(* Logix 5000 project; controller PLC_MCC1300_75F1 vendor 1 type 14 code 166 rev 32.11; software revision 32.04; part 62 of 83 *)
(* tags used below, declared in another part *)
   CONST_rgdDestMask : DINT[32];   // Destination Mask
   CONST_tPlant : UDT_PLANT_CONSTANTS;
   GP_TrackingSearchPlate : GP_TrackingSearchPlate;
   GP_TrackingValidateIndex : GP_TrackingValidateIndex;
   M315_M1_DR_R1 : AXIS_CIP_DRIVE;
   M315_xReqStopPrevConvForPos : BOOL;
   M315Popup : MAC_Popup_ZC[2];
   M315Popup_HMR : MAC_Popup_ZC_HMR[2];
   M315Popup_HMW : MAC_Popup_ZC_HMW[2];
   M315Popup_PlateFreeTimeout : TIMER;
   M315Popup_xDrivePosEnable : BOOL;
   TMP_d : DINT;
   TMP_dDiffPhotocellStartConv0 : DINT;
   TMP_dEndSearch0 : DINT;
   TMP_dEndSearch1 : DINT;
   TMP_dFixedSideOffsetBoth : DINT;
   TMP_dFixedSideOffsetConvoy : DINT;
   TMP_dFixedSideOffsetDW : DINT;
   TMP_dFixedSideOffsetUP : DINT;
   TMP_dHalfConveyorLength : DINT;
   TMP_dHalfPlateLength : DINT;
   TMP_dIndex : DINT;
   TMP_dStartSearch0 : DINT;
   TMP_dStartSearch1 : DINT;
   TMP_xALLForSideLeg : BOOL;
   TMP_xAllLiteToCullet : BOOL;
   TMP_xAtLeastOneForSideLeg : BOOL;
   TMP_xAtLeastOneToCullet : BOOL;
   TMP_xPosHead : BOOL;
   xAlwaysOFF : BOOL;
   xAlwaysON : BOOL;
   xDebugOFF : BOOL;
   Z300_BufferPlate : UDT_LINE_BUFFER_PLATE;
   Z300_Conveyor : UDT_StandConv[29];
   Z300_Conveyor_IN_MOTION : MAC_Conveyor_ZC_IN_MOTION[29];
   Z300_Conveyor_OUT_MOTION : MAC_Conveyor_ZC_OUT_MOTION[29];
   Z300_LineTracking : UDT_LINE_TRACKING;
   Z301 : MAC_Zone_ML;
(* MainProgram, continued *)

ROUTINE M315Popup1_Logic   (* ladder *)
   // #####_CONSTANTS_#####
   0: NOP();
   1: XIC(xAlwaysON)OTE(M315Popup[1].ST_xTunnelType);
   2: DIV(Z300_LineTracking.rgtTrkConv[28].dLengthConveyor,2,TMP_dHalfConveyorLength);
   3: MOV(Z300_LineTracking.rgtTrkConv[28].dStartPosition_cmm,M315Popup[1].AUX_dStartPosition_cmm)MOV(Z300_LineTracking.rgtTrkConv[28].dEndPosition_cmm,M315Popup[1].AUX_dEndPosition_cmm)MOV(1500,M315Popup[1].AUX_dReactionTime_ms)MOV(200000,M315Popup[1].AUX_dWindowSearch_cmm)MOV(Z300_Conveyor[28].AUX_rgdCurrentSpeed_mm_min[0],M315Popup[1].AUX_dSpeedConveyor_mm_min);
   // #####_MATCH_#####
   4: NOP();
   5: XIC(Z301.ST_xEnableControlError)OTE(M315Popup[1].ST_xEnableControlError);
   // #####_ALARMS_#####
   6: NOP();
   7: JSR(M315Popup1_Faults,0);
   // #####_HMI_LOGICS_#####
   8: NOP();
   9: XIC(xAlwaysON)OTE(M315Popup[1].ST_xExternalConditionToRise);
   10: XIC(xAlwaysON)OTE(M315Popup[1].ST_xExternalConditionToDescend);
   // #####_STATUSES_#####
   11: NOP();
   12: [XIC(M315Popup[1].ST_xStopMachineFault) ,XIC(M315Popup[1].ST_xStopNextCycleFault) ]OTE(M315Popup[1].ST_xMachineAlarm);
   13: [XIO(M315Popup[1].ST_xPhasesInProgress) ,XIO(M315Popup[1].ST_xOutputEnable) ]OTE(M315Popup[1].ST_xConditionOKForStopCycle);
   14: XIC(Z301.ST_xCycleON)XIO(M315Popup[1].ST_xManualMode)XIO(M315Popup[1].ST_xMachineAlarm)OTE(M315Popup[1].ST_xOutputEnable);
   15: XIC(Z301.ST_xCycleON)XIC(M315Popup[1].ST_xOutputEnable)XIO(M315Popup[1].ST_xPhasesInProgress)XIO(M315Popup[1].INPUT_xPopupHigh)XIC(M315Popup[1].INPUT_xPopupLow)XIO(M315Popup[1].ST_xCleaningAccepted)OTE(M315Popup[1].ST_xInitialConditionForRise);
   16: XIC(Z301.ST_xCycleON)XIC(M315Popup[1].ST_xOutputEnable)XIO(M315Popup[1].ST_xPhasesInProgress)XIO(M315Popup[1].INPUT_xPopupLow)XIC(M315Popup[1].INPUT_xPopupHigh)XIO(M315Popup[1].ST_xCleaningAccepted)OTE(M315Popup[1].ST_xInitialConditionForDescend);
   17: [XIC(M315Popup_HMW[1].xEnableDisableManualCommand) XIC(xAlwaysOFF) ,XIC(Z300_Conveyor[23].ST_xManualCmdEnabled) ]XIC(M315Popup[1].ST_xConditionOKForStopCycle)XIC(M315Popup[1].ST_xConditionOKForStopCycle)OTE(M315Popup[1].ST_xManualMode);
   18: XIO(M315Popup[1].ST_xManualMode)MOV(0,M315Popup_HMW[1].rgxMan);
   // #####_PHASES_&_LOGICS_#####
   19: NOP();
   20: XIC(xAlwaysON)OTE(M315Popup[1].ST_xCleaningConditionOK);
   21: [XIC(M315Popup_HMW[1].xLocalCleaningRequest) XIC(xAlwaysOFF) ,XIC(Z300_Conveyor[28].ST_xCleaningEnabled) XIC(M315Popup[1].INPUT_xPopupLow) ][XIC(M315Popup[1].ST_xCleaningConditionOK) ,XIC(M315Popup[1].ST_xCleaningAccepted) ]OTE(M315Popup[1].ST_xCleaningAccepted);
   22: XIC(M315Popup[1].ST_xInitialConditionForRise)XIC(M315Popup[1].ST_xExternalConditionToRise)XIC(M315Popup[1].ST_xRequestRise)XIO(M315Popup[1].PH_xRise)OTL(M315Popup[1].PH_xRise);
   23: XIC(M315Popup[1].PH_xRise)XIC(M315Popup[1].INPUT_xPopupHigh)XIO(M315Popup[1].INPUT_xPopupLow)[OTU(M315Popup[1].PH_xRise) ,OTE(M315Popup[1].PH_xEndRise) ];
   24: XIC(M315Popup[1].ST_xInitialConditionForDescend)XIC(M315Popup[1].ST_xExternalConditionToDescend)XIC(M315Popup[1].ST_xRequestDescend)[XIC(M315Popup[0].ST_xRequestDescend) ,XIC(M315Popup[0].INPUT_xPopupLow) ]XIO(M315Popup[1].PH_xDescend)OTL(M315Popup[1].PH_xDescend);
   25: XIC(M315Popup[1].PH_xDescend)XIC(M315Popup[1].INPUT_xPopupLow)XIO(M315Popup[1].INPUT_xPopupHigh)[OTU(M315Popup[1].PH_xDescend) ,OTE(M315Popup[1].PH_xEndDescend) ];
   26: [XIC(M315Popup[1].PH_xRise) ,XIC(M315Popup[1].PH_xEndRise) ,XIC(M315Popup[1].PH_xDescend) ,XIC(M315Popup[1].PH_xEndDescend) ]OTE(M315Popup[1].ST_xPhasesInProgress);
   27: [XIC(M315Popup[1].PH_xEndDescend) ,XIO(xAlwaysOFF) XIC(M315Popup[0].INPUT_xPopupLow) XIC(M315Popup[1].INPUT_xPopupLow) ]OTU(M315Popup[1].ST_xPlatePresence);
   28: XIO(M315Popup[1].ST_xPhasesInProgress)[XIC(M315Popup[1].INPUT_xPopupLow) XIO(M315Popup[1].INPUT_xPopupHigh) ,XIC(M315Popup[1].ST_xTunnelType) XIC(M315Popup[1].INPUT_xPopupHigh) XIO(M315Popup[1].INPUT_xPopupLow) ]OTE(M315Popup[1].ST_xOutOfEncumbrance);
   29: XIO(M315Popup[1].ST_xPhasesInProgress)XIO(M315Popup[1].ST_xPlatePresence)XIO(M315Popup[1].INPUT_xPopupHigh)XIC(M315Popup[1].INPUT_xPopupLow)OTE(M315Popup[1].ST_xConditionToReceiveGlass);
   30: XIO(M315Popup[1].ST_xPhasesInProgress)XIC(M315Popup[1].INPUT_xPopupHigh)XIO(M315Popup[1].INPUT_xPopupLow)OTE(M315Popup[1].ST_xConditionForUpperConveyor);
   // #####_EXTERNAL_DEVICE_#####
   31: NOP();
   // #####_HMI_STATUSES_#####
   32: NOP();
   33: XIC(M315Popup[1].INPUT_xPopupHigh)OTE(M315Popup_HMR[1].xHighPosition);
   34: XIC(M315Popup[1].INPUT_xPopupLow)OTE(M315Popup_HMR[1].xLowPosition);
   35: [MOV(1,M315Popup_HMR[1].rgdState) ,[XIC(M315Popup[1].OUTPUT_xPopupLifting) ,XIC(M315Popup[1].OUTPUT_xPopupDescent) ] MOV(3,M315Popup_HMR[1].rgdState) ,XIC(M315Popup[1].ST_xMachineWarning) MOV(5,M315Popup_HMR[1].rgdState) ,XIC(M315Popup[1].ST_xMachineAlarm) MOV(7,M315Popup_HMR[1].rgdState) ];
   36: XIC(M315Popup[1].ST_xCleaningAccepted)OTE(M315Popup_HMR[1].xPopUpCleaningEnabled);
   37: XIC(M315Popup[1].ST_xManualMode)XIC(M315Popup_HMW[1].rgxMan.0)XIC(M315Popup[1].OUTPUT_xPopupLifting)OTE(M315Popup_HMR[1].rgxMan.0);
   38: XIC(M315Popup[1].ST_xManualMode)XIC(M315Popup_HMW[1].rgxMan.1)XIC(M315Popup[1].OUTPUT_xPopupDescent)OTE(M315Popup_HMR[1].rgxMan.1);
   39: XIC(M315Popup[1].ST_xManualMode)XIC(M315Popup_HMW[1].rgxMan.8)XIC(M315Popup[1].OUTPUT_xRun)OTE(M315Popup_HMR[1].rgxMan.8);
   40: XIC(M315Popup[1].ST_xManualMode)XIC(M315Popup_HMW[1].rgxMan.9)XIC(M315Popup[1].OUTPUT_xReverse)OTE(M315Popup_HMR[1].rgxMan.9);
END_ROUTINE

ROUTINE M315PopupManagement   (* ladder *)
   // #####_CONSTANTS_#####
   0: NOP();
   1: MOV(CONST_rgdDestMask[2],M315Popup[0].AUX_dDestMaskOppOpSide)MOV(CONST_rgdDestMask[2],M315Popup[1].AUX_dDestMaskOppOpSide)MOV(20000,TMP_dFixedSideOffsetUP)MOV(-20000,TMP_dFixedSideOffsetDW)MOV(43000,TMP_dFixedSideOffsetBoth)MOV(30000,TMP_dFixedSideOffsetConvoy)MOV(380000,TMP_dHalfConveyorLength);
   // #####_MATCH_#####
   2: NOP();
   3: MOV(Z300_LineTracking.rgtTrkConv[26].dStartPosition_cmm,M315Popup[0].AUX_dStartPosition_cmm)MOV(Z300_LineTracking.rgtTrkConv[27].dEndPosition_cmm,M315Popup[0].AUX_dEndPosition_cmm)MOV(M315Popup[0].AUX_dEndPosition_cmm,M315Popup[1].AUX_dStartPosition_cmm)MOV(Z300_LineTracking.rgtTrkConv[28].dEndPosition_cmm,M315Popup[1].AUX_dEndPosition_cmm);
   4: MOV(Z300_LineTracking.rgtTrkConv[26].dStartPosition_cmm,M315Popup[0].AUX_dPosPhotocell_cmm)MOV(Z300_LineTracking.rgtTrkConv[26].dStartPosition_cmm,M315Popup[1].AUX_dPosPhotocell_cmm)SUB(Z300_LineTracking.rgtTrkConv[26].dStartPosition_cmm,M315Popup[0].AUX_dPosPhotocell_cmm,TMP_dDiffPhotocellStartConv0)MOV(50,M315Popup[0].tmOF_Wait.PRE)MOV(50,M315Popup[1].tmOF_Wait.PRE)MOV(10000,M315Popup[0].tmON_Saturation.PRE)MOV(10000,M315Popup[1].tmON_Saturation.PRE);
   5: SUB(M315Popup[0].AUX_dPosPhotocell_cmm,300000,TMP_dStartSearch0)SUB(M315Popup[0].AUX_dPosPhotocell_cmm,0,TMP_dEndSearch0)SUB(M315Popup[0].AUX_dPosPhotocell_cmm,300000,TMP_dStartSearch1)SUB(M315Popup[0].AUX_dPosPhotocell_cmm,0,TMP_dEndSearch1);
   // Set Positioning Type
   6: XIC(xAlwaysON)OTE(TMP_xPosHead);
   // ##### PREVIOUS CONVEYOR #####
   7: NOP();
   // Search plate limits
   8: MUL(M315Popup[0].AUX_dSpeedConveyor_mm_min,M315Popup[0].AUX_dReactionTime_ms,TMP_d)DIV(TMP_d,600,M315Popup[0].AUX_tSearchPlateData.dReaction_cmm);
   9: MOV(TMP_dStartSearch0,M315Popup[0].AUX_tSearchPlateData.dPositionDecision_cmm)MOV(TMP_dEndSearch0,M315Popup[0].AUX_tSearchPlateData.dPositionStopSearch_cmm)ADD(Z300_LineTracking.rgtTrkConv[28].dEndPosition_cmm,300000,M315Popup[0].AUX_tSearchPlateData.dPositionStopHooked_cmm);
   // Search plate on previous conveyor (reverse search)
   10: XIO(M315Popup[0].AUX_tSearchPlateData.xPlateHooked)GP_TrackingSearchPlate(GP_TrackingSearchPlate,M315Popup[0].AUX_tSearchPlateData.dPositionStopSearch_cmm,M315Popup[0].AUX_tSearchPlateData.dPositionDecision_cmm,0,Z300_LineTracking,M315Popup[0].AUX_tSearchPlateData.tResult,CONST_tPlant.dNumOfConveyors,CONST_tPlant.dNumCapsConveyor,Z300_BufferPlate);
   11: XIO(Z300_LineTracking.rgtTrkConv[25].xGlassPresence)XIO(Z300_LineTracking.rgtTrkConv[26].xGlassPresence)XIO(Z300_LineTracking.rgtTrkConv[27].xGlassPresence)XIO(Z300_LineTracking.rgtTrkConv[28].xGlassPresence)XIC(TMP_xPosHead)XIO(M315Popup[0].AUX_tSearchPlateData.tResult.xHeadPresence)MOV(0,M315Popup[0].AUX_tSearchPlateData.dIndex)MOV(0,M315Popup[0].AUX_dIndexHead);
   12: XIO(Z300_LineTracking.rgtTrkConv[25].xGlassPresence)XIO(Z300_LineTracking.rgtTrkConv[26].xGlassPresence)XIO(Z300_LineTracking.rgtTrkConv[27].xGlassPresence)XIO(Z300_LineTracking.rgtTrkConv[28].xGlassPresence)XIO(TMP_xPosHead)XIO(M315Popup[0].AUX_tSearchPlateData.tResult.xTailPresence)MOV(0,M315Popup[0].AUX_tSearchPlateData.dIndex)MOV(0,M315Popup[0].AUX_dIndexTail);
   13: XIC(TMP_xPosHead)XIC(M315Popup[0].AUX_tSearchPlateData.tResult.xHeadPresence)MOV(M315Popup[0].AUX_tSearchPlateData.tResult.rgdHeadPointer[0],M315Popup[0].AUX_dIndexHead);
   14: XIO(TMP_xPosHead)XIC(M315Popup[0].AUX_tSearchPlateData.tResult.xTailPresence)MOV(M315Popup[0].AUX_tSearchPlateData.tResult.rgdTailPointer[0],M315Popup[0].AUX_dIndexTail);
   15: XIO(M315Popup[0].AUX_tSearchPlateData.xPlateHooked)[XIC(TMP_xPosHead) XIC(M315Popup[0].AUX_tSearchPlateData.tResult.xHeadPresence) MOV(M315Popup[0].AUX_tSearchPlateData.tResult.rgdHeadPointer[0],M315Popup[0].AUX_tSearchPlateData.dIndex) ,XIO(TMP_xPosHead) XIC(M315Popup[0].AUX_tSearchPlateData.tResult.xTailPresence) MOV(M315Popup[0].AUX_tSearchPlateData.tResult.rgdTailPointer[0],M315Popup[0].AUX_tSearchPlateData.dIndex) ][OSR(M315Popup[0].AUX_tSearchPlateData.OSR_xPlateInWindows,M315Popup[0].AUX_tSearchPlateData.OS_xPlateInWindows) ,OSF(M315Popup[0].AUX_tSearchPlateData.OSF_xPlateInWindows,M315Popup[0].AUX_tSearchPlateData.OF_xPlateInWindows) ];
   16: GRT(M315Popup[0].AUX_tSearchPlateData.dIndex,0)[OTU(TMP_xAtLeastOneForSideLeg) ,OTL(TMP_xALLForSideLeg) ,OTL(TMP_xAllLiteToCullet) ,OTU(TMP_xAtLeastOneToCullet) ];
   // Verify destination
   17: GRT(M315Popup[0].AUX_tSearchPlateData.dIndex,0)JSR(sbrCheckConvoyZCDestination,5,M315Popup[0].AUX_tSearchPlateData.dIndex,M315Popup[0].AUX_dDestMaskOppOpSide,CONST_rgdDestMask[24],TMP_xAtLeastOneForSideLeg,TMP_xAllLiteToCullet,TMP_xAtLeastOneForSideLeg,TMP_xAllLiteToCullet)JSR(sbrCheckConvoyZCDestinationFull,5,M315Popup[0].AUX_tSearchPlateData.dIndex,M315Popup[0].AUX_dDestMaskOppOpSide,CONST_rgdDestMask[24],TMP_xALLForSideLeg,TMP_xAtLeastOneToCullet,TMP_xALLForSideLeg,TMP_xAtLeastOneToCullet)[XIC(TMP_xAtLeastOneForSideLeg) XIC(TMP_xALLForSideLeg) OTE(M315Popup[0].ST_xPlateComingToPopup) ,XIO(TMP_xALLForSideLeg) MOV(M315Popup[0].AUX_tSearchPlateData.dIndex,M315Popup[0].AUX_dIndexPlateFree) ];
   18: GP_TrackingValidateIndex(GP_TrackingValidateIndex,Z300_BufferPlate,M315Popup[0].AUX_tSearchPlateData.dIDMemory,M315Popup[0].AUX_tSearchPlateData.dIndex,M315Popup[0].AUX_tSearchPlateData.xIndexCons);
   // Check plate dimension
   19: XIC(M315Popup[0].ST_xPlateComingToPopup)MOV(M315Popup[0].AUX_tSearchPlateData.dIndex,TMP_dIndex)[LEQ(Z300_BufferPlate.rgtPlate[TMP_dIndex].tData.dTotalCaps,1) [GRT(Z300_BufferPlate.rgtPlate[TMP_dIndex].tData.dLength_cmm,TMP_dHalfConveyorLength) OTE(M315Popup[0].ST_xPlateToBothComing) ,XIO(M315Popup[0].ST_xPlateToBothComing) OTE(M315Popup[0].ST_xPlateToSingleComing) ] ,GRT(Z300_BufferPlate.rgtPlate[TMP_dIndex].tData.dTotalCaps,1) [LEQ(Z300_BufferPlate.rgtPlate[TMP_dIndex].tData.dLength_cmm,CONST_tPlant.rgdConvoyLimits_cmm[2]) ,XIO(xAlwaysOFF) ] OTE(M315Popup[0].ST_xConvoyComing) ];
   20: [XIC(Z300_Conveyor[25].xReqStop) ,XIO(xAlwaysOFF) ]XIC(M315Popup[0].ST_xPhasesInProgress)TOF(M315Popup[0].tmOF_Wait,?,?);
   21: [XIC(Z300_Conveyor[25].xReqStop) ,XIO(xAlwaysOFF) ]XIC(M315Popup[1].ST_xPhasesInProgress)TOF(M315Popup[1].tmOF_Wait,?,?);
   // Plate has left popup conveyors
   22: GRT(M315Popup[0].AUX_dIndexPlateFree,0)MOV(M315Popup[0].AUX_dIndexPlateFree,TMP_dIndex)GEQ(Z300_BufferPlate.rgtPlate[TMP_dIndex].tTracking.dPositionTail_cmm,Z300_LineTracking.rgtTrkConv[24].dEndPosition_cmm)MOV(0,M315Popup[0].AUX_dIndexPlateFree);
   // Stop previuos conveyor if no condition on pop-up conveyor
   23: [[XIC(M315Popup[0].ST_xPlateToSingleComing) [XIO(M315Popup[0].ST_xInitialConditionForRise) ,XIC(M315Popup[0].ST_xPlatePresentOnPopup) ,XIC(M315Popup[0].ST_xPlatePresence) ,XIC(Z300_LineTracking.rgtTrkConv[26].xGlassPresence) ,XIC(Z300_LineTracking.rgtTrkConv[27].xGlassPresence) ,EQU(M315Popup[0].AUX_dIndexPositioning,0) [XIC(M315Popup[0].ST_xPlateUnderPopup) ,XIC(M315Popup[1].ST_xPlateUnderPopup) ] ] ,XIC(M315Popup[0].ST_xPlateToSingleComing) [XIO(M315Popup[1].ST_xInitialConditionForRise) ,XIC(M315Popup[1].ST_xPlatePresentOnPopup) ,XIC(M315Popup[1].ST_xPlatePresence) ,XIC(Z300_LineTracking.rgtTrkConv[26].xGlassPresence) ,XIC(Z300_LineTracking.rgtTrkConv[27].xGlassPresence) ,XIC(Z300_LineTracking.rgtTrkConv[28].xGlassPresence) ,EQU(M315Popup[0].AUX_dIndexPositioning,0) [XIC(M315Popup[0].ST_xPlateUnderPopup) ,XIC(M315Popup[1].ST_xPlateUnderPopup) ] ] ,[XIC(M315Popup[0].ST_xPlateToBothComing) ,XIC(M315Popup[0].ST_xConvoyComing) ] [XIO(M315Popup[1].ST_xInitialConditionForRise) ,XIC(M315Popup[1].ST_xPlatePresentOnPopup) ,XIC(M315Popup[1].ST_xPlatePresence) ,XIC(Z300_LineTracking.rgtTrkConv[26].xGlassPresence) ,XIC(Z300_LineTracking.rgtTrkConv[27].xGlassPresence) ,XIC(Z300_LineTracking.rgtTrkConv[28].xGlassPresence) ,EQU(M315Popup[0].AUX_dIndexPositioning,0) XIC(M315Popup[1].ST_xPlateUnderPopup) ,XIO(M315Popup[0].ST_xInitialConditionForRise) ,XIC(M315Popup[0].ST_xPlatePresentOnPopup) ,XIC(M315Popup[0].ST_xPlatePresence) ,EQU(M315Popup[0].AUX_dIndexPositioning,0) XIC(M315Popup[0].ST_xPlateUnderPopup) ] ] ,XIO(M315Popup[0].INPUT_xPopupHigh) XIO(M315Popup[0].INPUT_xPopupLow) ,XIO(M315Popup[1].INPUT_xPopupHigh) XIO(M315Popup[1].INPUT_xPopupLow) ,XIC(M315_xReqStopPrevConvForPos) ,XIC(Z300_Conveyor[26].xReqExtStopLoadNewPlate) ,[XIC(M315Popup[0].ST_xPlateInPositionToRise) ,XIC(M315Popup[1].ST_xPlateInPositionToRise) ] ,XIC(Z300_Conveyor[26].ST_xCleaningEnabled) XIO(Z300_Conveyor[25].ST_xCleaningEnabled) ,XIC(M315Popup[0].ST_xPrevConvFreeAfterPos) ,XIC(M315Popup[1].ST_xPrevConvFreeAfterPos) ,[XIO(M315Popup[0].INPUT_xPopupHigh) ,XIO(M315Popup[1].INPUT_xPopupHigh) ] ,GRT(M315Popup[0].AUX_dIndexPositioning,0) [GRT(M315Popup[0].AUX_tSearchPlateData.dIndex,0) NEQ(M315Popup[0].AUX_tSearchPlateData.dIndex,M315Popup[0].AUX_dIndexPositioning) ,GRT(M315Popup[0].AUX_dIndexPlatePositioned,0) NEQ(M315Popup[0].AUX_dIndexPlatePositioned,M315Popup[0].AUX_dIndexPositioning) ] ,GRT(M315Popup[0].AUX_dIndexPlateFree,0) MOV(M315Popup[0].AUX_dIndexPlateFree,TMP_dIndex) [XIC(M315Popup[0].ST_xPlateToSingleComing) LES(Z300_BufferPlate.rgtPlate[TMP_dIndex].tTracking.dPositionTail_cmm,M315Popup[1].AUX_dStartPosition_cmm) ,[XIC(M315Popup[0].ST_xPlateToBothComing) ,XIC(M315Popup[0].ST_xConvoyComing) ,XIC(M315Popup[1].ST_xPlateToSingleComing) ] LES(Z300_BufferPlate.rgtPlate[TMP_dIndex].tTracking.dPositionTail_cmm,Z300_LineTracking.rgtTrkConv[24].dEndPosition_cmm) ] ]OTE(M315Popup[0].ST_xConditionToStopPrevious);
   24: XIO(xDebugOFF)GRT(M315Popup[0].AUX_dIndexPlateFree,0)XIC(Z300_Conveyor[26].ST_xRotationFeedback)MOV(10000,M315Popup_PlateFreeTimeout.PRE)[TON(M315Popup_PlateFreeTimeout,?,?) ,XIC(M315Popup_PlateFreeTimeout.DN) MOV(0,M315Popup[0].AUX_dIndexPlateFree) ];
   25: XIO(Z300_LineTracking.rgtTrkConv[26].xGlassPresence)XIO(Z300_LineTracking.rgtTrkConv[27].xGlassPresence)XIO(Z300_LineTracking.rgtTrkConv[28].xGlassPresence)XIC(Z300_Conveyor[26].ST_xRotationFeedback)XIC(Z300_Conveyor[27].ST_xRotationFeedback)XIC(Z300_Conveyor[28].ST_xRotationFeedback)[GRT(M315Popup[0].AUX_dIndexPlateFree,0) ,GRT(M315Popup[0].AUX_dIndexPlatePositioned,0) ]MOV(5000,M315Popup_PlateFreeTimeout.PRE)[TON(M315Popup_PlateFreeTimeout,?,?) ,XIC(M315Popup_PlateFreeTimeout.DN) [MOV(0,M315Popup[0].AUX_dIndexPlateFree) ,MOV(0,M315Popup[0].AUX_dIndexPlatePositioned) ] ];
   26: XIO(M315Popup[0].ST_xPlateUnderPopup)XIO(M315Popup[1].ST_xPlateUnderPopup)MOV(0,M315Popup[0].AUX_dIndexPlatePositioned);
   27: XIC(M315Popup[0].ST_xConditionToStopPrevious)GEQ(Z300_LineTracking.rgtTrkConv[25].dHeadPosition_cmm,Z300_Conveyor[25].AUX_rgdLoadPreset_cmm[0])[XIO(Z300_Conveyor[26].OUTPUT_xPositioning.0) XIO(M315Popup[0].tmON_Positioning.EN) ,[XIC(M315_xReqStopPrevConvForPos) ,XIC(Z300_Conveyor[26].xReqExtStopLoadNewPlate) ] ]OTE(M315Popup[0].ST_xStopPreviousConveyor);
   // STOP CONVEYOR M360
   28: XIC(M315Popup[0].ST_xStopPreviousConveyor)OTE(Z300_Conveyor[25].xReqStop);
   // #####_POSITIONING_#####
   29: NOP();
   // Hook plate for positioning
   30: XIC(M315Popup[0].ST_xPlateComingToPopup)[XIC(M315Popup[0].ST_xPlateToBothComing) XIO(Z300_LineTracking.rgtTrkConv[26].xGlassPresence) XIO(Z300_LineTracking.rgtTrkConv[27].xGlassPresence) XIO(Z300_LineTracking.rgtTrkConv[28].xGlassPresence) XIO(M315Popup[0].ST_xPlatePresentOnPopup) XIO(M315Popup[0].ST_xPlatePresence) XIO(M315Popup[1].ST_xPlatePresentOnPopup) XIO(M315Popup[1].ST_xPlatePresence) ,XIC(M315Popup[0].ST_xConvoyComing) XIO(Z300_LineTracking.rgtTrkConv[26].xGlassPresence) XIO(Z300_LineTracking.rgtTrkConv[27].xGlassPresence) XIO(Z300_LineTracking.rgtTrkConv[28].xGlassPresence) XIO(M315Popup[0].ST_xPlatePresentOnPopup) XIO(M315Popup[0].ST_xPlatePresence) XIO(M315Popup[1].ST_xPlatePresentOnPopup) XIO(M315Popup[1].ST_xPlatePresence) ,XIC(M315Popup[1].ST_xPlateToSingleComing) XIO(Z300_LineTracking.rgtTrkConv[26].xGlassPresence) XIO(Z300_LineTracking.rgtTrkConv[27].xGlassPresence) XIO(Z300_LineTracking.rgtTrkConv[28].xGlassPresence) XIO(M315Popup[1].ST_xPlatePresentOnPopup) XIO(M315Popup[1].ST_xPlatePresence) ,XIC(M315Popup[0].ST_xPlateToSingleComing) XIO(Z300_LineTracking.rgtTrkConv[26].xGlassPresence) XIO(Z300_LineTracking.rgtTrkConv[27].xGlassPresence) XIO(M315Popup[0].ST_xPlatePresentOnPopup) XIO(M315Popup[0].ST_xPlatePresence) ]XIO(M315Popup[0].AUX_tSearchPlateData.xPlateHooked)EQU(M315Popup[0].AUX_dIndexPositioning,0)GRT(M315Popup[0].AUX_tSearchPlateData.dIndex,0)XIC(M315Popup[0].AUX_tSearchPlateData.xIndexCons)MOV(M315Popup[0].AUX_tSearchPlateData.dIndex,TMP_dIndex)GRT(Z300_BufferPlate.rgtPlate[TMP_dIndex].tTracking.dPositionHead_cmm,M315Popup[0].AUX_tSearchPlateData.dPositionDecision_cmm)[XIO(Z300_Conveyor[25].xReqStop) ,XIO(xAlwaysOFF) ]XIO(Z300_Conveyor[26].OUTPUT_xPositioning.0)XIO(Z300_Conveyor[27].OUTPUT_xPositioning.0)XIO(Z300_Conveyor[28].OUTPUT_xPositioning.0)XIO(M315Popup[0].ST_xPlateInPositionToRise)XIO(M315Popup[1].ST_xPlateInPositionToRise)[OTL(M315Popup[0].AUX_tSearchPlateData.xPlateHooked) ,MOV(M315Popup[0].AUX_tSearchPlateData.dIndex,M315Popup[0].AUX_dIndexPositioning) ,JSR(sbrTrackingPositioningStart,2,M315Popup[0].AUX_dIndexPositioning,TMP_xPosHead) ];
   31: GP_TrackingValidateIndex(GP_TrackingValidateIndex,Z300_BufferPlate,M315Popup[0].AUX_dMemoryPositioning,M315Popup[0].AUX_dIndexPositioning,M315Popup[0].ST_xIndexConsPositioning);
   // Check plate dimension
   32: XIC(M315Popup[0].AUX_tSearchPlateData.xPlateHooked)[XIC(M315Popup[0].ST_xIndexConsPositioning) ,XIO(xDebugOFF) ]XIO(M315Popup[0].ST_xPlateToBothPositioning)XIO(M315Popup[0].ST_xPlateToSinglePositioning)XIO(M315Popup[1].ST_xPlateToSinglePositioning)XIO(M315Popup[0].ST_xConvoyPositioning)MOV(M315Popup[0].AUX_dIndexPositioning,TMP_dIndex)[LEQ(Z300_BufferPlate.rgtPlate[TMP_dIndex].tData.dTotalCaps,1) [GRT(Z300_BufferPlate.rgtPlate[TMP_dIndex].tData.dLength_cmm,TMP_dHalfConveyorLength) OTL(M315Popup[0].ST_xPlateToBothPositioning) ,XIO(M315Popup[0].ST_xPlateToBothPositioning) OTL(M315Popup[0].ST_xPlateToSinglePositioning) ] ,GRT(Z300_BufferPlate.rgtPlate[TMP_dIndex].tData.dTotalCaps,1) [LEQ(Z300_BufferPlate.rgtPlate[TMP_dIndex].tData.dLength_cmm,CONST_tPlant.rgdConvoyLimits_cmm[2]) ,XIO(xAlwaysOFF) ] OTL(M315Popup[0].ST_xConvoyPositioning) ];
   // Positioning request (In case of head positioning also previous conveyors are involved)
   33: XIO(M315Popup[0].ST_xPlateInPositionToRise)XIO(M315Popup[1].ST_xPlateInPositionToRise)XIC(M315Popup[0].AUX_tSearchPlateData.xPlateHooked)[XIC(M315Popup[0].ST_xPlateToSinglePositioning) XIO(Z300_LineTracking.rgtTrkConv[26].xGlassPresence) XIO(Z300_LineTracking.rgtTrkConv[27].xGlassPresence) XIO(M315Popup[0].ST_xPlatePresence) [XIO(M315Popup[0].ST_xPlateUnderPopup) ,XIO(xDebugOFF) ] XIC(M315Popup[0].ST_xOutputEnable) XIC(M315Popup[0].INPUT_xPopupLow) XIC(M315Popup[0].ST_xInitialConditionForRise) ,XIC(M315Popup[1].ST_xPlateToSinglePositioning) XIO(Z300_LineTracking.rgtTrkConv[26].xGlassPresence) XIO(Z300_LineTracking.rgtTrkConv[27].xGlassPresence) XIO(Z300_LineTracking.rgtTrkConv[28].xGlassPresence) XIO(M315Popup[1].ST_xPlatePresence) XIO(M315Popup[0].ST_xPlateUnderPopup) [XIO(M315Popup[1].ST_xPlateUnderPopup) ,XIO(xDebugOFF) ] XIC(M315Popup[1].ST_xOutputEnable) XIC(M315Popup[1].INPUT_xPopupLow) XIC(M315Popup[1].ST_xInitialConditionForRise) ,XIC(M315Popup[0].ST_xPlateToBothPositioning) XIO(Z300_LineTracking.rgtTrkConv[26].xGlassPresence) XIO(Z300_LineTracking.rgtTrkConv[27].xGlassPresence) XIO(Z300_LineTracking.rgtTrkConv[28].xGlassPresence) XIO(M315Popup[0].ST_xPlatePresence) XIO(M315Popup[0].ST_xPlateUnderPopup) XIC(M315Popup[0].ST_xOutputEnable) XIC(M315Popup[0].INPUT_xPopupLow) XIC(M315Popup[0].ST_xInitialConditionForRise) XIO(M315Popup[1].ST_xPlatePresence) [XIO(M315Popup[1].ST_xPlateUnderPopup) ,XIO(xDebugOFF) ] XIC(M315Popup[1].ST_xOutputEnable) XIC(M315Popup[1].INPUT_xPopupLow) XIC(M315Popup[1].ST_xInitialConditionForRise) ,XIC(M315Popup[0].ST_xConvoyPositioning) XIO(Z300_LineTracking.rgtTrkConv[26].xGlassPresence) XIO(Z300_LineTracking.rgtTrkConv[27].xGlassPresence) XIO(Z300_LineTracking.rgtTrkConv[28].xGlassPresence) XIO(M315Popup[0].ST_xPlatePresence) XIO(M315Popup[0].ST_xPlateUnderPopup) XIC(M315Popup[0].ST_xOutputEnable) XIC(M315Popup[0].INPUT_xPopupLow) XIC(M315Popup[0].ST_xInitialConditionForRise) XIO(M315Popup[1].ST_xPlatePresence) [XIO(M315Popup[1].ST_xPlateUnderPopup) ,XIO(xDebugOFF) ] XIC(M315Popup[1].ST_xOutputEnable) XIC(M315Popup[1].INPUT_xPopupLow) XIC(M315Popup[1].ST_xInitialConditionForRise) ]XIO(Z300_Conveyor[26].xReqStop)XIO(Z300_Conveyor[27].xReqStop)[XIC(M315Popup[0].ST_xIndexConsPositioning) ,XIO(xDebugOFF) ][XIC(TMP_xPosHead) XIC(M315Popup[0].AUX_tSearchPlateData.tResult.xHeadPresence) ,XIO(TMP_xPosHead) XIC(M315Popup[0].AUX_tSearchPlateData.tResult.xTailPresence) ]XIO(Z300_Conveyor[26].xReqPositioningHead)XIO(Z300_Conveyor[26].xReqPositioningTail)XIO(Z300_Conveyor[27].xReqPositioningHead)XIO(Z300_Conveyor[27].xReqPositioningTail)[XIO(Z300_Conveyor[28].xReqStop) XIO(Z300_Conveyor[28].xReqPositioningHead) XIO(Z300_Conveyor[28].xReqPositioningTail) ,XIC(M315Popup[1].ST_xPlateToSinglePositioning) ]XIO(M315Popup[0].tmOF_Wait.DN)XIO(M315Popup[1].tmOF_Wait.DN)TON(M315Popup[0].tmON_Positioning,?,?)XIC(M315Popup[0].tmON_Positioning.DN)[XIC(TMP_xPosHead) [OTL(Z300_Conveyor[26].xReqPositioningHead) ,OTL(Z300_Conveyor[27].xReqPositioningHead) ] ,XIO(TMP_xPosHead) [OTL(Z300_Conveyor[26].xReqPositioningTail) ,OTL(Z300_Conveyor[27].xReqPositioningTail) ] ,OTE(M315Popup[0].OS_xStartPositioning) ,[XIC(M315Popup[0].ST_xPlateToBothPositioning) ,XIC(M315Popup[0].ST_xConvoyPositioning) ,XIC(M315Popup[1].ST_xPlateToSinglePositioning) ] [XIC(TMP_xPosHead) OTL(Z300_Conveyor[28].xReqPositioningHead) ,XIO(TMP_xPosHead) OTL(Z300_Conveyor[28].xReqPositioningTail) ,OTE(M315Popup[1].OS_xStartPositioning) ] ,OTU(Z300_Conveyor_OUT_MOTION[26].DR_MAR_M[0].PC) ,OTU(Z300_Conveyor_IN_MOTION[26].DR_MAR_M[0].PC) ,OTU(Z300_Conveyor_OUT_MOTION[27].DR_MAR_M[0].PC) ,OTU(Z300_Conveyor_IN_MOTION[27].DR_MAR_M[0].PC) ,OTU(Z300_Conveyor_OUT_MOTION[28].DR_MAR_M[0].PC) ,OTU(Z300_Conveyor_IN_MOTION[28].DR_MAR_M[0].PC) ,OTU(Z300_Conveyor_OUT_MOTION[26].DR_MAM_M[0].PC) ,OTU(Z300_Conveyor_IN_MOTION[26].DR_MAM_M[0].PC) ,OTU(Z300_Conveyor_OUT_MOTION[27].DR_MAM_M[0].PC) ,OTU(Z300_Conveyor_IN_MOTION[27].DR_MAM_M[0].PC) ,OTU(Z300_Conveyor_OUT_MOTION[28].DR_MAM_M[0].PC) ,OTU(Z300_Conveyor_IN_MOTION[28].DR_MAM_M[0].PC) ];
   // Target calculation
   34: [XIC(M315Popup[0].OS_xStartPositioning) ,XIC(M315Popup[1].OS_xStartPositioning) ][XIC(M315Popup[0].ST_xIndexConsPositioning) ,XIO(xDebugOFF) ]MOV(M315Popup[0].AUX_tSearchPlateData.dIndex,TMP_dIndex)[XIC(M315Popup[0].ST_xPlateToSinglePositioning) ADD(TMP_dDiffPhotocellStartConv0,TMP_dFixedSideOffsetUP,TMP_d) [XIC(TMP_xPosHead) ADD(TMP_d,TMP_dHalfConveyorLength,M315Popup[0].AUX_dReqTarget_cmm) GRT(Z300_BufferPlate.rgtPlate[TMP_dIndex].tData.dLength_cmm,335000) ADD(M315Popup[0].AUX_dReqTarget_cmm,15000,M315Popup[0].AUX_dReqTarget_cmm) ,XIO(TMP_xPosHead) ADD(TMP_d,Z300_BufferPlate.rgtPlate[TMP_dIndex].tData.dLength_cmm,M315Popup[0].AUX_dReqTarget_cmm) ] ,XIC(M315Popup[0].ST_xPlateToBothPositioning) DIV(Z300_BufferPlate.rgtPlate[TMP_dIndex].tData.dLength_cmm,2,TMP_dHalfPlateLength) ADD(TMP_dDiffPhotocellStartConv0,TMP_dHalfConveyorLength,TMP_d) ADD(TMP_d,TMP_dFixedSideOffsetBoth,TMP_d) [XIC(TMP_xPosHead) ADD(TMP_d,TMP_dHalfPlateLength,M315Popup[0].AUX_dReqTarget_cmm) ,XIO(TMP_xPosHead) SUB(TMP_d,TMP_dHalfPlateLength,M315Popup[0].AUX_dReqTarget_cmm) ] ,XIC(M315Popup[0].ST_xConvoyPositioning) DIV(Z300_BufferPlate.rgtPlate[TMP_dIndex].tData.rgtCap[0].dConvTotLength_cmm,2,TMP_dHalfPlateLength) ADD(TMP_dDiffPhotocellStartConv0,TMP_dHalfConveyorLength,TMP_d) ADD(TMP_d,TMP_dFixedSideOffsetConvoy,TMP_d) [XIC(TMP_xPosHead) ADD(TMP_d,TMP_dHalfPlateLength,M315Popup[0].AUX_dReqTarget_cmm) ,XIO(TMP_xPosHead) SUB(TMP_d,TMP_dHalfPlateLength,M315Popup[0].AUX_dReqTarget_cmm) ] ];
   // Final drive target (In case of head positioning also previous conveyors are involved)
   35: [XIC(M315Popup[0].OS_xStartPositioning) ,XIC(M315Popup[1].OS_xStartPositioning) ][XIC(M315Popup[0].ST_xIndexConsPositioning) ,XIO(xDebugOFF) ]SUB(M315Popup[0].AUX_dReqTarget_cmm,TMP_dDiffPhotocellStartConv0,TMP_d)ADD(TMP_d,Z300_LineTracking.rgtTrkConv[23].dStartPosition_cmm,TMP_d)ADD(TMP_d,150000,M315Popup[0].AUX_dPosTimeout)[[XIC(M315Popup[0].ST_xPlateToSinglePositioning) ,XIC(M315Popup[0].ST_xPlateToBothPositioning) ] ADD(M315Popup[0].AUX_dReqTarget_cmm,M315Popup_HMW[0].dSingleCapOffset_cmm,Z300_Conveyor[23].AUX_rgdTarget_cmm[0]) ,XIC(M315Popup[0].ST_xConvoyPositioning) ADD(M315Popup[0].AUX_dReqTarget_cmm,M315Popup_HMW[0].dConvoyOffset_cmm,Z300_Conveyor[23].AUX_rgdTarget_cmm[0]) ]XIC(TMP_xPosHead)[MOV(Z300_Conveyor[23].AUX_rgdTarget_cmm[0],Z300_Conveyor[22].AUX_rgdTarget_cmm[0]) ,XIO(M315Popup[0].ST_xPlateToSinglePositioning) MOV(Z300_Conveyor[23].AUX_rgdTarget_cmm[0],Z300_Conveyor[24].AUX_rgdTarget_cmm[1]) ];
   36: XIO(xDebugOFF)MOV(M315Popup[0].AUX_dIndexPositioning,TMP_dIndex)GRT(TMP_dIndex,0)LES(Z300_BufferPlate.rgtPlate[TMP_dIndex].tData.dTotalCaps,2)[XIC(Z300_Conveyor[26].OUTPUT_xPositioning.0) GEQ(Z300_BufferPlate.rgtPlate[TMP_dIndex].tTracking.dPositionHead_cmm,M315Popup[0].AUX_dStartPosition_cmm) XIO(M315_M1_DR_R1.Registration1InputStatus) XIC(M315Popup_xDrivePosEnable) ,XIC(Z300_Conveyor[26].xReqExtStopLoadNewPlate) ]OTE(Z300_Conveyor[26].xReqExtStopLoadNewPlate);
